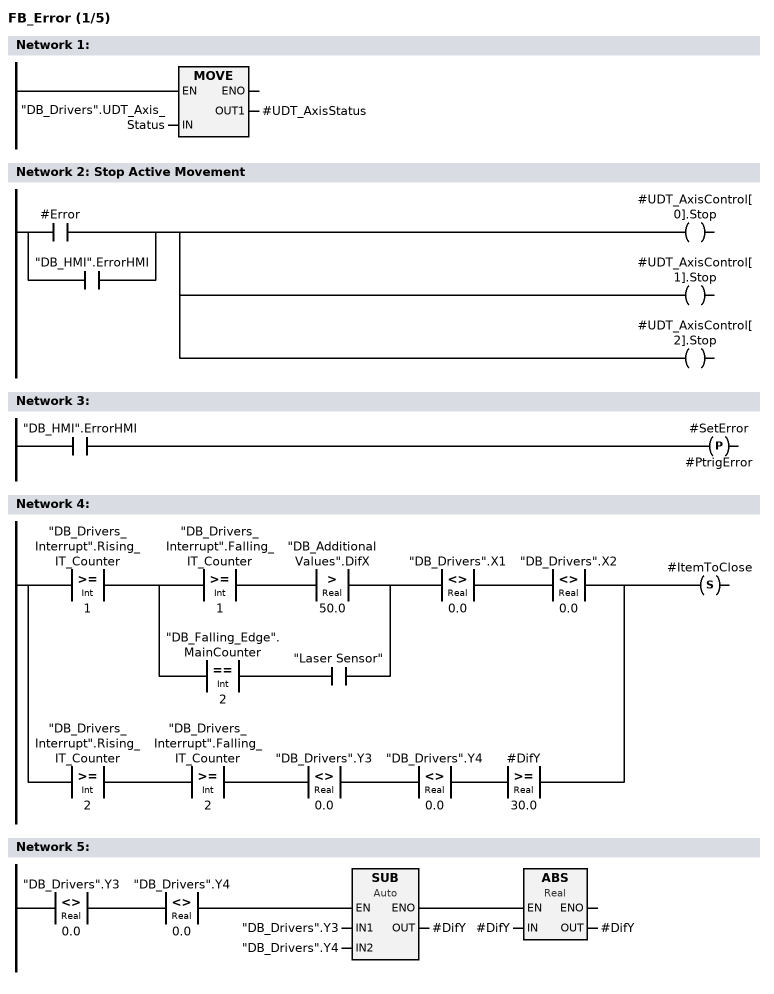
   RUNG wire#powerrail
      Move(in := "DB_Drivers".UDT_Axis_Status, out1 => #UDT_AxisStatus)
   END_RUNG
   // the same network as SCL:
   #UDT_AxisStatus := "DB_Drivers".UDT_Axis_Status;
END_REGION

REGION Network 2: Stop Active Movement
   RUNG wire#powerrail
      Contact( #Error )
      wire#w1
      Coil( #UDT_AxisControl[0].Stop )
   END_RUNG
   RUNG wire#powerrail
      Contact( "DB_HMI".ErrorHMI )
   END_RUNG wire#w1
   RUNG wire#w1
      Coil( #UDT_AxisControl[1].Stop )
   END_RUNG
   RUNG wire#w1
      Coil( #UDT_AxisControl[2].Stop )
   END_RUNG
   // the same network as SCL:
   #UDT_AxisControl[0].Stop := #Error OR "DB_HMI".ErrorHMI;
   #UDT_AxisControl[1].Stop := #Error OR "DB_HMI".ErrorHMI;
   #UDT_AxisControl[2].Stop := #Error OR "DB_HMI".ErrorHMI;
END_REGION

REGION Network 3
   #SetError := "DB_HMI".ErrorHMI AND NOT #PtrigError;   // rising edge
   #PtrigError := "DB_HMI".ErrorHMI;
END_REGION

REGION Network 4
   RUNG wire#powerrail
      { S7_Templates := "SrcType := Int" } GE_Contact(in1 := "DB_Drivers_Interrupt".Rising_IT_Counter, in2 := 1)
      wire#w1
      { S7_Templates := "SrcType := Int" } GE_Contact(in1 := "DB_Drivers_Interrupt".Falling_IT_Counter, in2 := 1)
      { S7_Templates := "SrcType := Real" } GT_Contact(in1 := "DB_AdditionalValues".DifX, in2 := 50.0)
      wire#w2
      { S7_Templates := "SrcType := Real" } NE_Contact(in1 := "DB_Drivers".X1, in2 := 0.0)
      { S7_Templates := "SrcType := Real" } NE_Contact(in1 := "DB_Drivers".X2, in2 := 0.0)
      wire#w3
      S_Coil( #ItemToClose )
   END_RUNG
   RUNG wire#w1
      { S7_Templates := "SrcType := Int" } EQ_Contact(in1 := "DB_Falling_Edge".MainCounter, in2 := 2)
      Contact( "Laser Sensor" )
   END_RUNG wire#w2
   RUNG wire#powerrail
      { S7_Templates := "SrcType := Int" } GE_Contact(in1 := "DB_Drivers_Interrupt".Rising_IT_Counter, in2 := 2)
      { S7_Templates := "SrcType := Int" } GE_Contact(in1 := "DB_Drivers_Interrupt".Falling_IT_Counter, in2 := 2)
      { S7_Templates := "SrcType := Real" } NE_Contact(in1 := "DB_Drivers".Y3, in2 := 0.0)
      { S7_Templates := "SrcType := Real" } NE_Contact(in1 := "DB_Drivers".Y4, in2 := 0.0)
      { S7_Templates := "SrcType := Real" } GE_Contact(in1 := #DifY, in2 := 30.0)
   END_RUNG wire#w3
   // the same network as SCL:
   IF (("DB_Drivers_Interrupt".Rising_IT_Counter >= 1) AND ((("DB_Drivers_Interrupt".Falling_IT_Counter >= 1) AND ("DB_AdditionalValues".DifX > 50.0)) OR (("DB_Falling_Edge".MainCounter = 2) AND "Laser Sensor")) AND ("DB_Drivers".X1 <> 0.0) AND ("DB_Drivers".X2 <> 0.0)) OR (("DB_Drivers_Interrupt".Rising_IT_Counter >= 2) AND ("DB_Drivers_Interrupt".Falling_IT_Counter >= 2) AND ("DB_Drivers".Y3 <> 0.0) AND ("DB_Drivers".Y4 <> 0.0) AND (#DifY >= 30.0)) THEN
       #ItemToClose := TRUE;
   END_IF;
END_REGION

REGION Network 5
   RUNG wire#powerrail
      { S7_Templates := "SrcType := Real" } NE_Contact(in1 := "DB_Drivers".Y3, in2 := 0.0)
      { S7_Templates := "SrcType := Real" } NE_Contact(in1 := "DB_Drivers".Y4, in2 := 0.0)
      Sub(in1 := "DB_Drivers".Y3, in2 := "DB_Drivers".Y4, out => #DifY)
      { S7_Templates := "SrcType := Real" } Abs(in := #DifY, out => #DifY)
   END_RUNG
   // the same network as SCL:
   IF ("DB_Drivers".Y3 <> 0.0) AND ("DB_Drivers".Y4 <> 0.0) THEN
       #DifY := "DB_Drivers".Y3 - "DB_Drivers".Y4;
       #DifY := ABS(#DifY);
   END_IF;
END_REGION

REGION Network 6
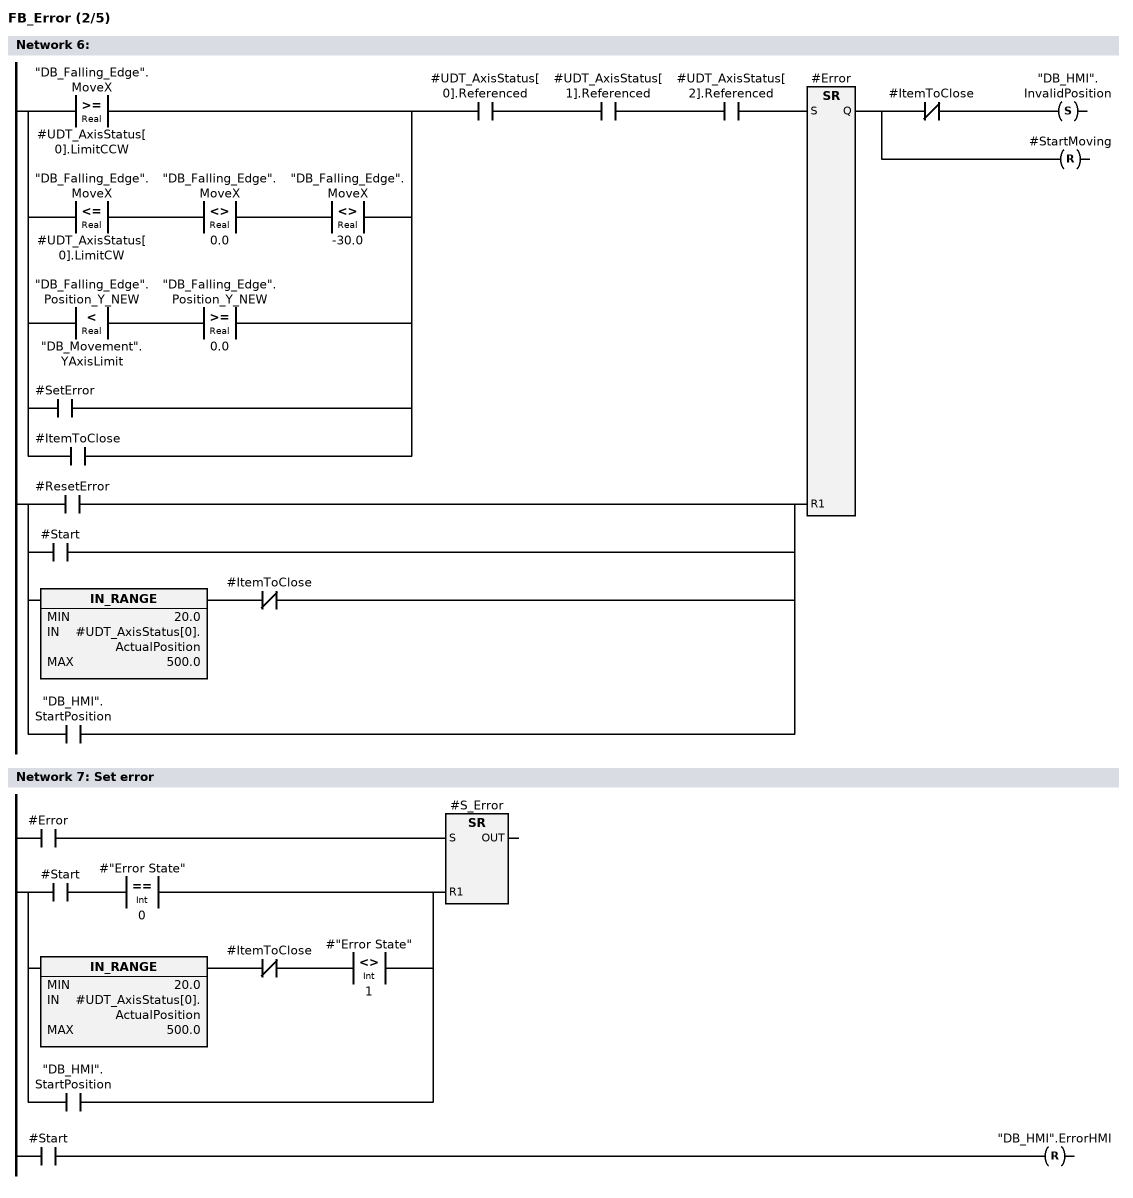
   RUNG wire#powerrail
      { S7_Templates := "SrcType := Real" } GE_Contact(in1 := "DB_Falling_Edge".MoveX, in2 := #UDT_AxisStatus[0].LimitCCW)
      wire#w1
      Contact( #UDT_AxisStatus[0].Referenced )
      Contact( #UDT_AxisStatus[1].Referenced )
      Contact( #UDT_AxisStatus[2].Referenced )
      S_SR(operand := #Error, r1 := wire#w2)
      wire#w3
      I_Contact( #ItemToClose )
      S_Coil( "DB_HMI".InvalidPosition )
   END_RUNG
   RUNG wire#powerrail
      { S7_Templates := "SrcType := Real" } LE_Contact(in1 := "DB_Falling_Edge".MoveX, in2 := #UDT_AxisStatus[0].LimitCW)
      { S7_Templates := "SrcType := Real" } NE_Contact(in1 := "DB_Falling_Edge".MoveX, in2 := 0.0)
      { S7_Templates := "SrcType := Real" } NE_Contact(in1 := "DB_Falling_Edge".MoveX, in2 := -30.0)
   END_RUNG wire#w1
   RUNG wire#powerrail
      { S7_Templates := "SrcType := Real" } LT_Contact(in1 := "DB_Falling_Edge".Position_Y_NEW, in2 := "DB_Movement".YAxisLimit)
      { S7_Templates := "SrcType := Real" } GE_Contact(in1 := "DB_Falling_Edge".Position_Y_NEW, in2 := 0.0)
   END_RUNG wire#w1
   RUNG wire#powerrail
      Contact( #SetError )
   END_RUNG wire#w1
   RUNG wire#powerrail
      Contact( #ItemToClose )
   END_RUNG wire#w1
   RUNG wire#powerrail
      Contact( #ResetError )
   END_RUNG wire#w2
   RUNG wire#powerrail
      Contact( #Start )
   END_RUNG wire#w2
   RUNG wire#powerrail
      { S7_Templates := "SrcType := Real" } InRange(min := 20.0, in := #UDT_AxisStatus[0].ActualPosition, max := 500.0)
      I_Contact( #ItemToClose )
   END_RUNG wire#w2
   RUNG wire#powerrail
      Contact( "DB_HMI".StartPosition )
   END_RUNG wire#w2
   RUNG wire#w3
      R_Coil( #StartMoving )
   END_RUNG
   // the same network as SCL:
   IF (("DB_Falling_Edge".MoveX >= #UDT_AxisStatus[0].LimitCCW) OR (("DB_Falling_Edge".MoveX <= #UDT_AxisStatus[0].LimitCW) AND ("DB_Falling_Edge".MoveX <> 0.0) AND ("DB_Falling_Edge".MoveX <> (-30.0))) OR (("DB_Falling_Edge".Position_Y_NEW < "DB_Movement".YAxisLimit) AND ("DB_Falling_Edge".Position_Y_NEW >= 0.0)) OR #SetError OR #ItemToClose) AND #UDT_AxisStatus[0].Referenced AND #UDT_AxisStatus[1].Referenced AND #UDT_AxisStatus[2].Referenced THEN
       #Error := TRUE;   // SR flip-flop
   END_IF;
   IF #ResetError OR #Start OR ((20.0 <= #UDT_AxisStatus[0].ActualPosition) AND (#UDT_AxisStatus[0].ActualPosition <= 500.0) AND NOT #ItemToClose) OR "DB_HMI".StartPosition THEN
       #Error := FALSE;
   END_IF;
   IF #Error AND NOT #ItemToClose THEN "DB_HMI".InvalidPosition := TRUE; END_IF;
   IF #Error THEN #StartMoving := FALSE; END_IF;
END_REGION

REGION Network 7: Set error
   RUNG wire#powerrail
      Contact( #Error )
      S_SR(operand := #S_Error, r1 := wire#w1)
   END_RUNG
   RUNG wire#powerrail
      Contact( #Start )
      { S7_Templates := "SrcType := Int" } EQ_Contact(in1 := #"Error State", in2 := 0)
   END_RUNG wire#w1
   RUNG wire#powerrail
      { S7_Templates := "SrcType := Real" } InRange(min := 20.0, in := #UDT_AxisStatus[0].ActualPosition, max := 500.0)
      I_Contact( #ItemToClose )
      { S7_Templates := "SrcType := Int" } NE_Contact(in1 := #"Error State", in2 := 1)
   END_RUNG wire#w1
   RUNG wire#powerrail
      Contact( "DB_HMI".StartPosition )
   END_RUNG wire#w1
   RUNG wire#powerrail
      Contact( #Start )
      R_Coil( "DB_HMI".ErrorHMI )
   END_RUNG
   // the same network as SCL:
   IF #Error THEN
       #S_Error := TRUE;   // SR flip-flop
   END_IF;
   IF (#Start AND (#"Error State" = 0)) OR ((20.0 <= #UDT_AxisStatus[0].ActualPosition) AND (#UDT_AxisStatus[0].ActualPosition <= 500.0) AND NOT #ItemToClose AND (#"Error State" <> 1)) OR "DB_HMI".StartPosition THEN
       #S_Error := FALSE;
   END_IF;
   IF #Start THEN "DB_HMI".ErrorHMI := FALSE; END_IF;
END_REGION

REGION Network 8: Set color of error ind
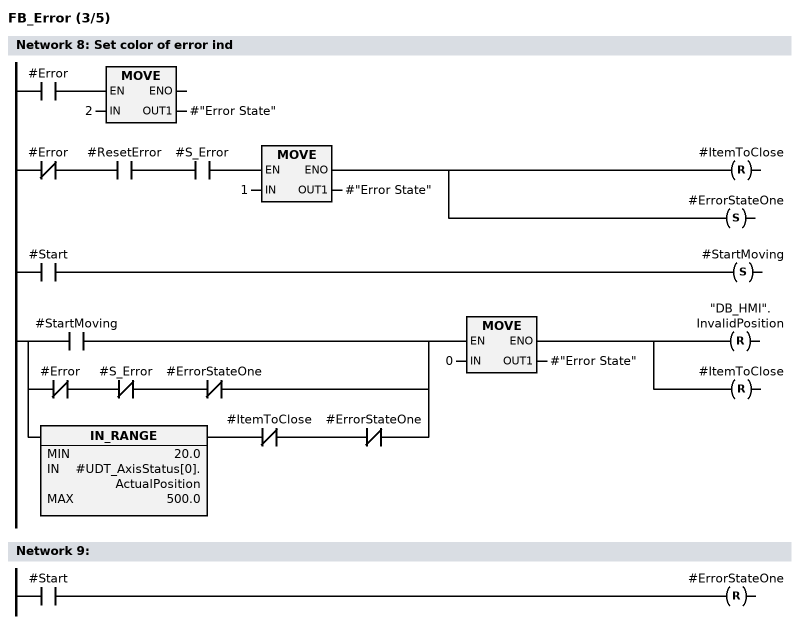
   RUNG wire#powerrail
      Contact( #Error )
      Move(in := 2, out1 => #"Error State")
   END_RUNG
   RUNG wire#powerrail
      I_Contact( #Error )
      Contact( #ResetError )
      Contact( #S_Error )
      Move(in := 1, out1 => #"Error State")
      wire#w1
      R_Coil( #ItemToClose )
   END_RUNG
   RUNG wire#w1
      S_Coil( #ErrorStateOne )
   END_RUNG
   RUNG wire#powerrail
      Contact( #Start )
      S_Coil( #StartMoving )
   END_RUNG
   RUNG wire#powerrail
      Contact( #StartMoving )
      wire#w2
      Move(in := 0, out1 => #"Error State")
      wire#w3
      R_Coil( "DB_HMI".InvalidPosition )
   END_RUNG
   RUNG wire#powerrail
      I_Contact( #Error )
      I_Contact( #S_Error )
      I_Contact( #ErrorStateOne )
   END_RUNG wire#w2
   RUNG wire#powerrail
      { S7_Templates := "SrcType := Real" } InRange(min := 20.0, in := #UDT_AxisStatus[0].ActualPosition, max := 500.0)
      I_Contact( #ItemToClose )
      I_Contact( #ErrorStateOne )
   END_RUNG wire#w2
   RUNG wire#w3
      R_Coil( #ItemToClose )
   END_RUNG
   // the same network as SCL:
   IF #Error THEN #"Error State" := 2; END_IF;
   IF NOT #Error AND #ResetError AND #S_Error THEN
       #"Error State" := 1;
       #ItemToClose := FALSE;
       #ErrorStateOne := TRUE;
   END_IF;
   IF #Start THEN #StartMoving := TRUE; END_IF;
   IF #StartMoving OR (NOT #Error AND NOT #S_Error AND NOT #ErrorStateOne) OR ((20.0 <= #UDT_AxisStatus[0].ActualPosition) AND (#UDT_AxisStatus[0].ActualPosition <= 500.0) AND NOT #ItemToClose AND NOT #ErrorStateOne) THEN
       #"Error State" := 0;
       "DB_HMI".InvalidPosition := FALSE;
       #ItemToClose := FALSE;
   END_IF;
END_REGION

REGION Network 9
   RUNG wire#powerrail
      Contact( #Start )
      R_Coil( #ErrorStateOne )
   END_RUNG
   // the same network as SCL:
   IF #Start THEN #ErrorStateOne := FALSE; END_IF;
END_REGION

REGION Network 10: Reset error
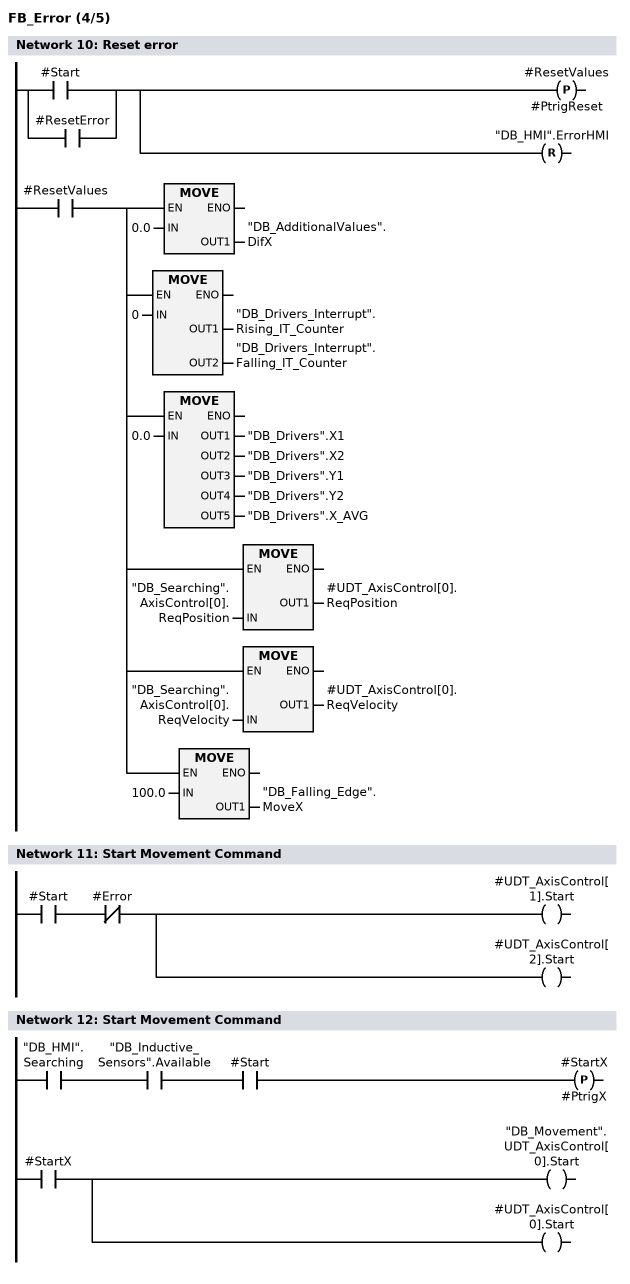
   #_w1 := #Start OR #ResetError;
   #ResetValues := #_w1 AND NOT #PtrigReset;   // rising edge
   #PtrigReset := #_w1;
   IF #_w1 THEN "DB_HMI".ErrorHMI := FALSE; END_IF;
   IF #ResetValues THEN
       "DB_AdditionalValues".DifX := 0.0;
       "DB_Drivers_Interrupt".Rising_IT_Counter := 0;
       "DB_Drivers_Interrupt".Falling_IT_Counter := 0;
       "DB_Drivers".X1 := 0.0;
       "DB_Drivers".X2 := 0.0;
       "DB_Drivers".Y1 := 0.0;
       "DB_Drivers".Y2 := 0.0;
       "DB_Drivers".X_AVG := 0.0;
       #UDT_AxisControl[0].ReqPosition := "DB_Searching".AxisControl[0].ReqPosition;
       #UDT_AxisControl[0].ReqVelocity := "DB_Searching".AxisControl[0].ReqVelocity;
       "DB_Falling_Edge".MoveX := 100.0;
   END_IF;
END_REGION

REGION Network 11: Start Movement Command
   RUNG wire#powerrail
      Contact( #Start )
      I_Contact( #Error )
      wire#w1
      Coil( #UDT_AxisControl[1].Start )
   END_RUNG
   RUNG wire#w1
      Coil( #UDT_AxisControl[2].Start )
   END_RUNG
   // the same network as SCL:
   #UDT_AxisControl[1].Start := #Start AND NOT #Error;
   #UDT_AxisControl[2].Start := #Start AND NOT #Error;
END_REGION

REGION Network 12: Start Movement Command
   #_w1 := "DB_HMI".Searching AND "DB_Inductive_Sensors".Available AND #Start;
   #StartX := #_w1 AND NOT #PtrigX;   // rising edge
   #PtrigX := #_w1;
   "DB_Movement".UDT_AxisControl[0].Start := #StartX;
   #UDT_AxisControl[0].Start := #StartX;
END_REGION

REGION Network 13: Active error
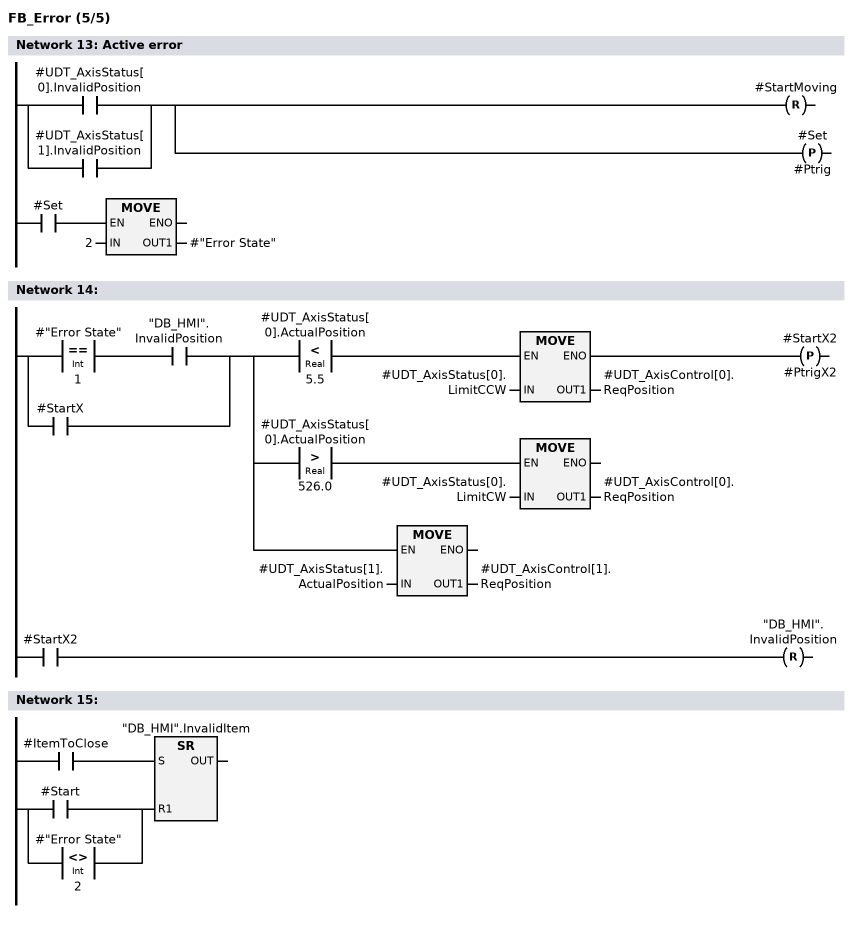
   #_w1 := #UDT_AxisStatus[0].InvalidPosition OR #UDT_AxisStatus[1].InvalidPosition;
   IF #_w1 THEN #StartMoving := FALSE; END_IF;
   #Set := #_w1 AND NOT #Ptrig;   // rising edge
   #Ptrig := #_w1;
   IF #Set THEN #"Error State" := 2; END_IF;
END_REGION

REGION Network 14
   #_w1 := ((#"Error State" = 1) AND "DB_HMI".InvalidPosition) OR #StartX;
   #_w2 := #_w1 AND (#UDT_AxisStatus[0].ActualPosition < 5.5);
   IF #_w2 THEN #UDT_AxisControl[0].ReqPosition := #UDT_AxisStatus[0].LimitCCW; END_IF;
   #StartX2 := #_w2 AND NOT #PtrigX2;   // rising edge
   #PtrigX2 := #_w2;
   IF #_w1 AND (#UDT_AxisStatus[0].ActualPosition > 526.0) THEN
       #UDT_AxisControl[0].ReqPosition := #UDT_AxisStatus[0].LimitCW;
   END_IF;
   IF #_w1 THEN #UDT_AxisControl[1].ReqPosition := #UDT_AxisStatus[1].ActualPosition; END_IF;
   IF #StartX2 THEN "DB_HMI".InvalidPosition := FALSE; END_IF;
END_REGION

REGION Network 15
   RUNG wire#powerrail
      Contact( #ItemToClose )
      S_SR(operand := "DB_HMI".InvalidItem, r1 := wire#w1)
   END_RUNG
   RUNG wire#powerrail
      Contact( #Start )
   END_RUNG wire#w1
   RUNG wire#powerrail
      { S7_Templates := "SrcType := Int" } NE_Contact(in1 := #"Error State", in2 := 2)
   END_RUNG wire#w1
   // the same network as SCL:
   IF #ItemToClose THEN
       "DB_HMI".InvalidItem := TRUE;   // SR flip-flop
   END_IF;
   IF #Start OR (#"Error State" <> 2) THEN "DB_HMI".InvalidItem := FALSE; END_IF;
END_REGION
END_FUNCTION_BLOCK

// folder: HMI

FUNCTION "FC_HMI" : Void   // FC2, LAD
TITLE = HMI interface
{ S7_Optimized_Access := 'TRUE' }
VERSION : 0.1
   VAR_TEMP
      StartPositionReached : Bool;
      PtrigSP : Bool;
   END_VAR
   VAR_TEMP   // added for the SCL form of the ladder/FBD networks
      _w1 : Bool;
   END_VAR
BEGIN

REGION Network 1: Center Position Counting
   // Set Actual Status: Center Position Counting
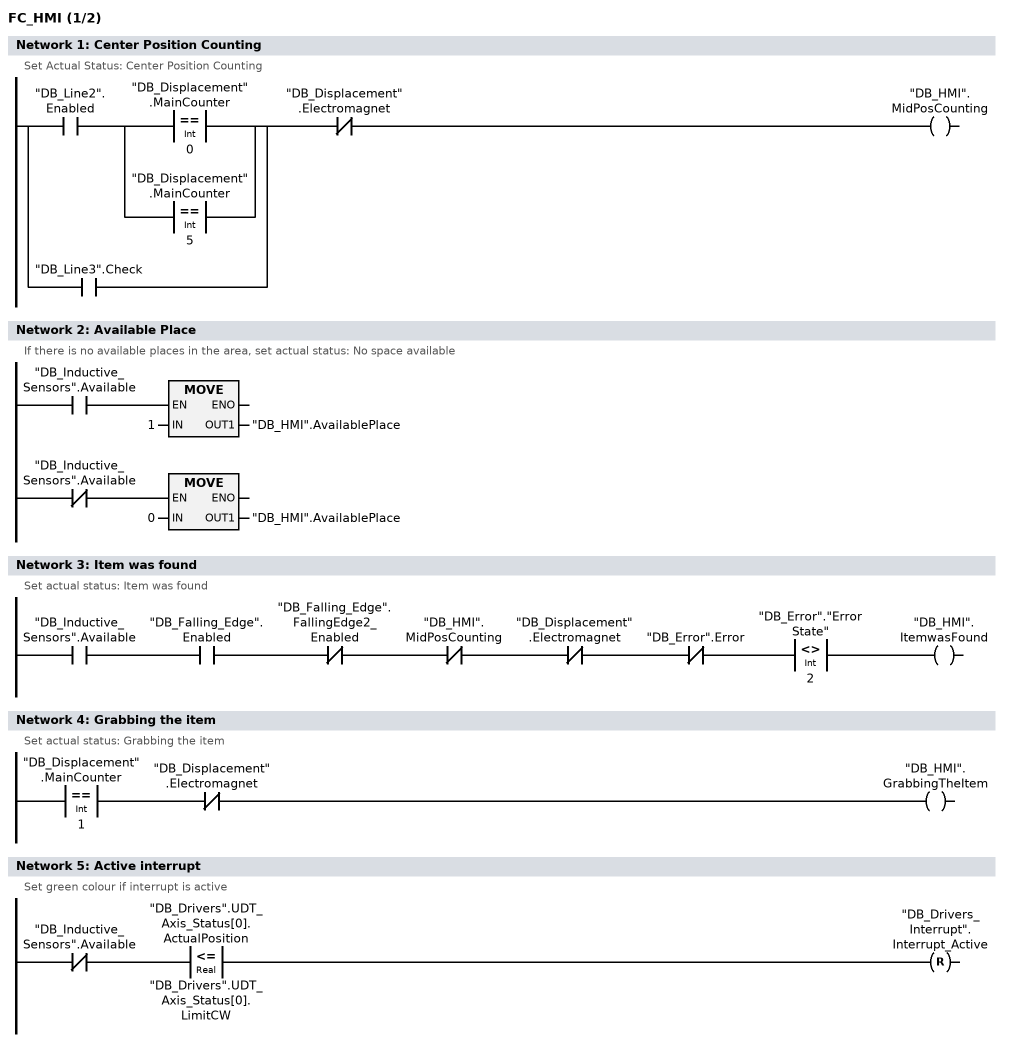
   RUNG wire#powerrail
      Contact( "DB_Line2".Enabled )
      wire#w1
      { S7_Templates := "SrcType := Int" } EQ_Contact(in1 := "DB_Displacement".MainCounter, in2 := 0)
      wire#w2
      I_Contact( "DB_Displacement".Electromagnet )
      Coil( "DB_HMI".MidPosCounting )
   END_RUNG
   RUNG wire#w1
      { S7_Templates := "SrcType := Int" } EQ_Contact(in1 := "DB_Displacement".MainCounter, in2 := 5)
   END_RUNG wire#w2
   RUNG wire#powerrail
      Contact( "DB_Line3".Check )
   END_RUNG wire#w2
   // the same network as SCL:
   "DB_HMI".MidPosCounting := (("DB_Line2".Enabled AND (("DB_Displacement".MainCounter = 0) OR ("DB_Displacement".MainCounter = 5))) OR "DB_Line3".Check) AND NOT "DB_Displacement".Electromagnet;
END_REGION

REGION Network 2: Available Place
   // If there is no available places in the area, set actual status: No space available
   RUNG wire#powerrail
      Contact( "DB_Inductive_Sensors".Available )
      Move(in := 1, out1 => "DB_HMI".AvailablePlace)
   END_RUNG
   RUNG wire#powerrail
      I_Contact( "DB_Inductive_Sensors".Available )
      Move(in := 0, out1 => "DB_HMI".AvailablePlace)
   END_RUNG
   // the same network as SCL:
   IF "DB_Inductive_Sensors".Available THEN "DB_HMI".AvailablePlace := 1; END_IF;
   IF NOT "DB_Inductive_Sensors".Available THEN "DB_HMI".AvailablePlace := 0; END_IF;
END_REGION

REGION Network 3: Item was found
   // Set actual status: Item was found
   RUNG wire#powerrail
      Contact( "DB_Inductive_Sensors".Available )
      Contact( "DB_Falling_Edge".Enabled )
      I_Contact( "DB_Falling_Edge".FallingEdge2_Enabled )
      I_Contact( "DB_HMI".MidPosCounting )
      I_Contact( "DB_Displacement".Electromagnet )
      I_Contact( "DB_Error".Error )
      { S7_Templates := "SrcType := Int" } NE_Contact(in1 := "DB_Error"."Error State", in2 := 2)
      Coil( "DB_HMI".ItemwasFound )
   END_RUNG
   // the same network as SCL:
   "DB_HMI".ItemwasFound := "DB_Inductive_Sensors".Available AND "DB_Falling_Edge".Enabled AND NOT "DB_Falling_Edge".FallingEdge2_Enabled AND NOT "DB_HMI".MidPosCounting AND NOT "DB_Displacement".Electromagnet AND NOT "DB_Error".Error AND ("DB_Error"."Error State" <> 2);
END_REGION

REGION Network 4: Grabbing the item
   // Set actual status: Grabbing the item
   RUNG wire#powerrail
      { S7_Templates := "SrcType := Int" } EQ_Contact(in1 := "DB_Displacement".MainCounter, in2 := 1)
      I_Contact( "DB_Displacement".Electromagnet )
      Coil( "DB_HMI".GrabbingTheItem )
   END_RUNG
   // the same network as SCL:
   "DB_HMI".GrabbingTheItem := ("DB_Displacement".MainCounter = 1) AND NOT "DB_Displacement".Electromagnet;
END_REGION

REGION Network 5: Active interrupt
   // Set green colour if interrupt is active
   RUNG wire#powerrail
      I_Contact( "DB_Inductive_Sensors".Available )
      { S7_Templates := "SrcType := Real" } LE_Contact(in1 := "DB_Drivers".UDT_Axis_Status[0].ActualPosition, in2 := "DB_Drivers".UDT_Axis_Status[0].LimitCW)
      R_Coil( "DB_Drivers_Interrupt".Interrupt_Active )
   END_RUNG
   // the same network as SCL:
   IF NOT "DB_Inductive_Sensors".Available AND ("DB_Drivers".UDT_Axis_Status[0].ActualPosition <= "DB_Drivers".UDT_Axis_Status[0].LimitCW) THEN
       "DB_Drivers_Interrupt".Interrupt_Active := FALSE;
   END_IF;
END_REGION

REGION Network 6: Start Position Reached
   // If 'Start position' button was pressed, set suitable status
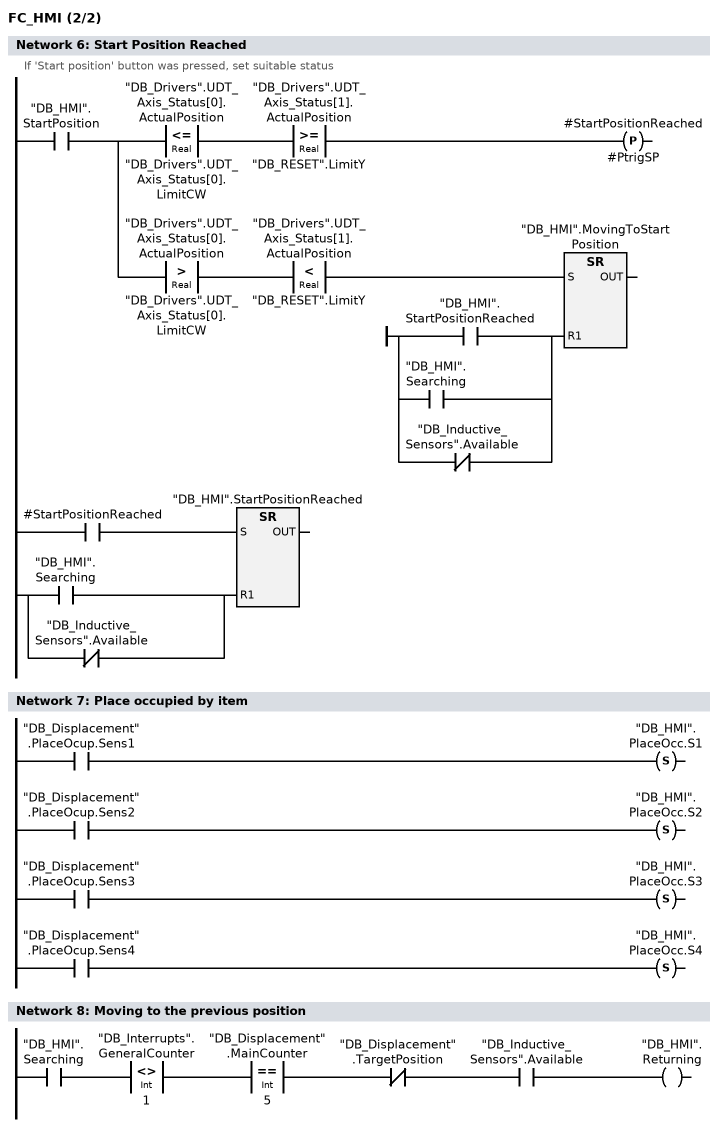
   #_w1 := "DB_HMI".StartPosition AND ("DB_Drivers".UDT_Axis_Status[0].ActualPosition <= "DB_Drivers".UDT_Axis_Status[0].LimitCW) AND ("DB_Drivers".UDT_Axis_Status[1].ActualPosition >= "DB_RESET".LimitY);
   #StartPositionReached := #_w1 AND NOT #PtrigSP;   // rising edge
   #PtrigSP := #_w1;
   IF "DB_HMI".StartPosition AND ("DB_Drivers".UDT_Axis_Status[0].ActualPosition > "DB_Drivers".UDT_Axis_Status[0].LimitCW) AND ("DB_Drivers".UDT_Axis_Status[1].ActualPosition < "DB_RESET".LimitY) THEN
       "DB_HMI".MovingToStartPosition := TRUE;   // SR flip-flop
   END_IF;
   IF "DB_HMI".StartPositionReached OR "DB_HMI".Searching OR NOT "DB_Inductive_Sensors".Available THEN
       "DB_HMI".MovingToStartPosition := FALSE;
   END_IF;
   IF #StartPositionReached THEN
       "DB_HMI".StartPositionReached := TRUE;   // SR flip-flop
   END_IF;
   IF "DB_HMI".Searching OR NOT "DB_Inductive_Sensors".Available THEN
       "DB_HMI".StartPositionReached := FALSE;
   END_IF;
END_REGION

REGION Network 7: Place occupied by item
   RUNG wire#powerrail
      Contact( "DB_Displacement".PlaceOcup.Sens1 )
      S_Coil( "DB_HMI".PlaceOcc.S1 )
   END_RUNG
   RUNG wire#powerrail
      Contact( "DB_Displacement".PlaceOcup.Sens2 )
      S_Coil( "DB_HMI".PlaceOcc.S2 )
   END_RUNG
   RUNG wire#powerrail
      Contact( "DB_Displacement".PlaceOcup.Sens3 )
      S_Coil( "DB_HMI".PlaceOcc.S3 )
   END_RUNG
   RUNG wire#powerrail
      Contact( "DB_Displacement".PlaceOcup.Sens4 )
      S_Coil( "DB_HMI".PlaceOcc.S4 )
   END_RUNG
   // the same network as SCL:
   IF "DB_Displacement".PlaceOcup.Sens1 THEN "DB_HMI".PlaceOcc.S1 := TRUE; END_IF;
   IF "DB_Displacement".PlaceOcup.Sens2 THEN "DB_HMI".PlaceOcc.S2 := TRUE; END_IF;
   IF "DB_Displacement".PlaceOcup.Sens3 THEN "DB_HMI".PlaceOcc.S3 := TRUE; END_IF;
   IF "DB_Displacement".PlaceOcup.Sens4 THEN "DB_HMI".PlaceOcc.S4 := TRUE; END_IF;
END_REGION

REGION Network 8: Moving to the previous position
   RUNG wire#powerrail
      Contact( "DB_HMI".Searching )
      { S7_Templates := "SrcType := Int" } NE_Contact(in1 := "DB_Interrupts".GeneralCounter, in2 := 1)
      { S7_Templates := "SrcType := Int" } EQ_Contact(in1 := "DB_Displacement".MainCounter, in2 := 5)
      I_Contact( "DB_Displacement".TargetPosition )
      Contact( "DB_Inductive_Sensors".Available )
      Coil( "DB_HMI".Returning )
   END_RUNG
   // the same network as SCL:
   "DB_HMI".Returning := "DB_HMI".Searching AND ("DB_Interrupts".GeneralCounter <> 1) AND ("DB_Displacement".MainCounter = 5) AND NOT "DB_Displacement".TargetPosition AND "DB_Inductive_Sensors".Available;
END_REGION
END_FUNCTION

// folder: OB

ORGANIZATION_BLOCK "Main"   // OB1, LAD, ProgramCycle
TITLE = "Main Program Sweep (Cycle)"
{ S7_Optimized_Access := 'TRUE' }
VERSION : 0.1
   VAR_INPUT
      Initial_Call : Bool;   // Initial call of this OB
      Remanence : Bool;   // =True, if remanent data are available
   END_VAR
BEGIN

REGION Network 1: Drivers Parameters
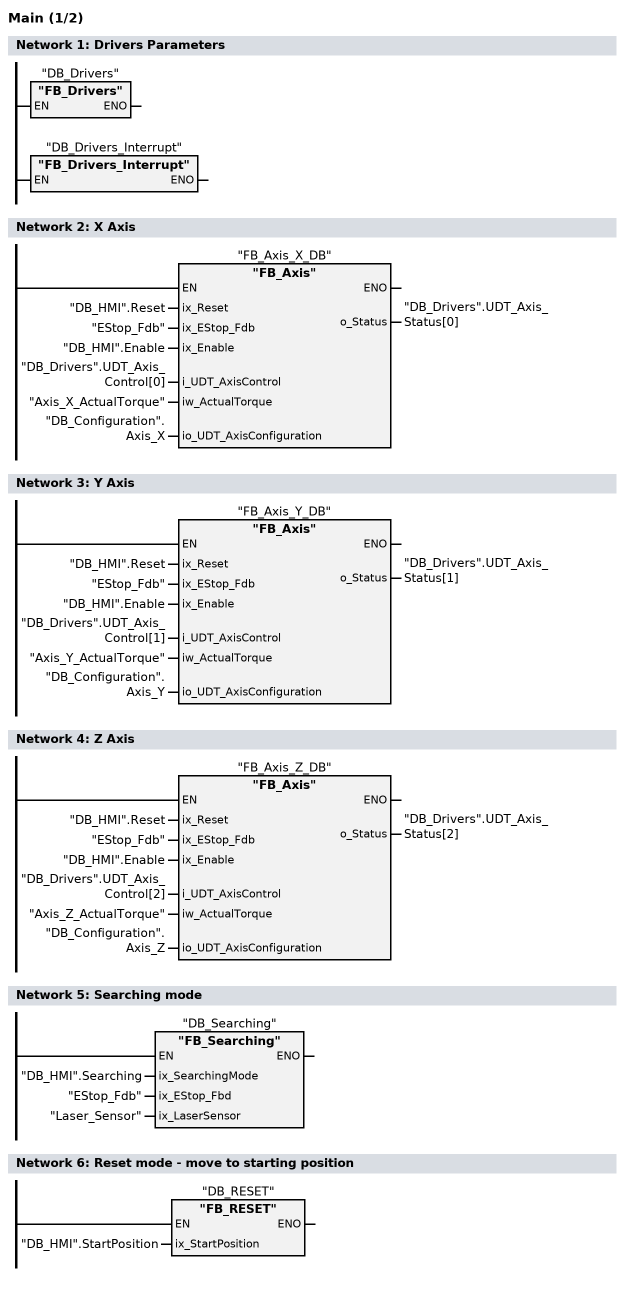
   RUNG wire#powerrail
      "DB_Drivers"()
   END_RUNG
   RUNG wire#powerrail
      "DB_Drivers_Interrupt"()
   END_RUNG
   // the same network as SCL:
   "DB_Drivers"();   // "FB_Drivers"
   "DB_Drivers_Interrupt"();   // "FB_Drivers_Interrupt"
END_REGION

REGION Network 2: X Axis
   RUNG wire#powerrail
      "FB_Axis_X_DB"(ix_Reset := "DB_HMI".Reset, ix_EStop_Fdb := "EStop_Fdb", ix_Enable := "DB_HMI".Enable, i_UDT_AxisControl := "DB_Drivers".UDT_Axis_Control[0], iw_ActualTorque := "Axis_X_ActualTorque", io_UDT_AxisConfiguration := "DB_Configuration".Axis_X, o_Status => "DB_Drivers".UDT_Axis_Status[0])
   END_RUNG
   // the same network as SCL:
   "FB_Axis_X_DB"(ix_Reset := "DB_HMI".Reset,   // "FB_Axis"
                  ix_EStop_Fdb := "EStop_Fdb",
                  ix_Enable := "DB_HMI".Enable,
                  i_UDT_AxisControl := "DB_Drivers".UDT_Axis_Control[0],
                  iw_ActualTorque := "Axis_X_ActualTorque",
                  io_UDT_AxisConfiguration := "DB_Configuration".Axis_X,
                  o_Status => "DB_Drivers".UDT_Axis_Status[0]);
END_REGION

REGION Network 3: Y Axis
   RUNG wire#powerrail
      "FB_Axis_Y_DB"(ix_Reset := "DB_HMI".Reset, ix_EStop_Fdb := "EStop_Fdb", ix_Enable := "DB_HMI".Enable, i_UDT_AxisControl := "DB_Drivers".UDT_Axis_Control[1], iw_ActualTorque := "Axis_Y_ActualTorque", io_UDT_AxisConfiguration := "DB_Configuration".Axis_Y, o_Status => "DB_Drivers".UDT_Axis_Status[1])
   END_RUNG
   // the same network as SCL:
   "FB_Axis_Y_DB"(ix_Reset := "DB_HMI".Reset,   // "FB_Axis"
                  ix_EStop_Fdb := "EStop_Fdb",
                  ix_Enable := "DB_HMI".Enable,
                  i_UDT_AxisControl := "DB_Drivers".UDT_Axis_Control[1],
                  iw_ActualTorque := "Axis_Y_ActualTorque",
                  io_UDT_AxisConfiguration := "DB_Configuration".Axis_Y,
                  o_Status => "DB_Drivers".UDT_Axis_Status[1]);
END_REGION

REGION Network 4: Z Axis
   RUNG wire#powerrail
      "FB_Axis_Z_DB"(ix_Reset := "DB_HMI".Reset, ix_EStop_Fdb := "EStop_Fdb", ix_Enable := "DB_HMI".Enable, i_UDT_AxisControl := "DB_Drivers".UDT_Axis_Control[2], iw_ActualTorque := "Axis_Z_ActualTorque", io_UDT_AxisConfiguration := "DB_Configuration".Axis_Z, o_Status => "DB_Drivers".UDT_Axis_Status[2])
   END_RUNG
   // the same network as SCL:
   "FB_Axis_Z_DB"(ix_Reset := "DB_HMI".Reset,   // "FB_Axis"
                  ix_EStop_Fdb := "EStop_Fdb",
                  ix_Enable := "DB_HMI".Enable,
                  i_UDT_AxisControl := "DB_Drivers".UDT_Axis_Control[2],
                  iw_ActualTorque := "Axis_Z_ActualTorque",
                  io_UDT_AxisConfiguration := "DB_Configuration".Axis_Z,
                  o_Status => "DB_Drivers".UDT_Axis_Status[2]);
END_REGION

REGION Network 5: Searching mode
   RUNG wire#powerrail
      "DB_Searching"(ix_SearchingMode := "DB_HMI".Searching, ix_EStop_Fbd := "EStop_Fdb", ix_LaserSensor := "Laser_Sensor")
   END_RUNG
   // the same network as SCL:
   "DB_Searching"(ix_SearchingMode := "DB_HMI".Searching,   // "FB_Searching"
                  ix_EStop_Fbd := "EStop_Fdb",
                  ix_LaserSensor := "Laser_Sensor");
END_REGION

REGION Network 6: Reset mode - move to starting position
   RUNG wire#powerrail
      "DB_RESET"(ix_StartPosition := "DB_HMI".StartPosition)
   END_RUNG
   // the same network as SCL:
   "DB_RESET"(ix_StartPosition := "DB_HMI".StartPosition);   // "FB_RESET"
END_REGION

REGION Network 7: Interrupt Function 1
